REGION Network 9
   RUNG wire#powerrail
      Contact( "I1_7" )
      wire#w1
      Contact( "DB12"."2#回转窑烟气管道闸板上升" )
      I_Contact( "I1_5" )
      I_Contact( "闸阀上限" )
      I_Contact( "Q2_1" )
      Coil( "Q2_0" )
   END_RUNG
   RUNG wire#w1
      Contact( "DB12"."2#回转窑烟气管道闸板下降" )
      I_Contact( "I1_6" )
      I_Contact( "闸阀下限" )
      I_Contact( "Q2_0" )
      Coil( "Q2_1" )
   END_RUNG
   // the same network as SCL:
   "Q2_0" := "I1_7" AND "DB12"."2#回转窑烟气管道闸板上升" AND NOT "I1_5" AND NOT "闸阀上限" AND NOT "Q2_1";
   "Q2_1" := "I1_7" AND "DB12"."2#回转窑烟气管道闸板下降" AND NOT "I1_6" AND NOT "闸阀下限" AND NOT "Q2_0";
END_REGION

REGION Network 10
   RUNG wire#powerrail
      Contact( "DB22".STAT3 )
      Contact( "尾排风机高压远程" )
      Coil( "尾排风机高压合闸驱动" )
   END_RUNG
   // the same network as SCL:
   "尾排风机高压合闸驱动" := "DB22".STAT3 AND "尾排风机高压远程";
END_REGION

REGION Network 11
   RUNG wire#powerrail
      Contact( "DB22".STAT4 )
      Coil( "尾排风机高压分闸驱动" )
   END_RUNG
   // the same network as SCL:
   "尾排风机高压分闸驱动" := "DB22".STAT4;
END_REGION

REGION Network 12
   RUNG wire#powerrail
      Contact( "DB22".STAT5 )
      wire#w1
      Contact( "尾排风机变频远程" )
      Contact( "尾排风机变频待机" )
      I_Contact( "尾排风机变频故障" )
      wire#w2
      I_Contact( "Tag_24" )
      Coil( "尾排风机高压柜变频启动" )
   END_RUNG
   RUNG wire#powerrail
      Contact( "尾排风机高压柜变频启动" )
   END_RUNG wire#w1
   RUNG wire#w2
      S_ODT(T_NO := "Tag_24", TV := S5T#3S, R :=, BI =>, RET_VAL =>)
   END_RUNG
   // the same network as SCL:
   #_w1 := ("DB22".STAT5 OR "尾排风机高压柜变频启动") AND "尾排风机变频远程" AND "尾排风机变频待机" AND NOT "尾排风机变频故障";
   "尾排风机高压柜变频启动" := #_w1 AND NOT "Tag_24";
   #_s5time1 := S_ODT(T_NO := "Tag_24", S := #_w1, TV := S5T#3S);
END_REGION

REGION Network 13
   RUNG wire#powerrail
      Contact( "DB22".STAT6 )
      wire#w1
      Contact( "尾排风机变频远程" )
      wire#w2
      I_Contact( "Tag_25" )
      Coil( "尾排风机高压柜变频停止" )
   END_RUNG
   RUNG wire#powerrail
      Contact( "尾排风机变频故障" )
   END_RUNG wire#w1
   RUNG wire#powerrail
      Contact( "尾排风机高压柜变频停止" )
   END_RUNG wire#w1
   RUNG wire#w2
      S_ODT(T_NO := "Tag_25", TV := S5T#3S, R :=, BI =>, RET_VAL =>)
   END_RUNG
   // the same network as SCL:
   #_w1 := ("DB22".STAT6 OR "尾排风机变频故障" OR "尾排风机高压柜变频停止") AND "尾排风机变频远程";
   "尾排风机高压柜变频停止" := #_w1 AND NOT "Tag_25";
   #_s5time1 := S_ODT(T_NO := "Tag_25", S := #_w1, TV := S5T#3S);
END_REGION
END_FUNCTION

FUNCTION "回转窑模拟量给定" : Void   // FC14, LAD
{ S7_Optimized_Access := 'FALSE' }
VERSION : 0.1
BEGIN

REGION Network 1
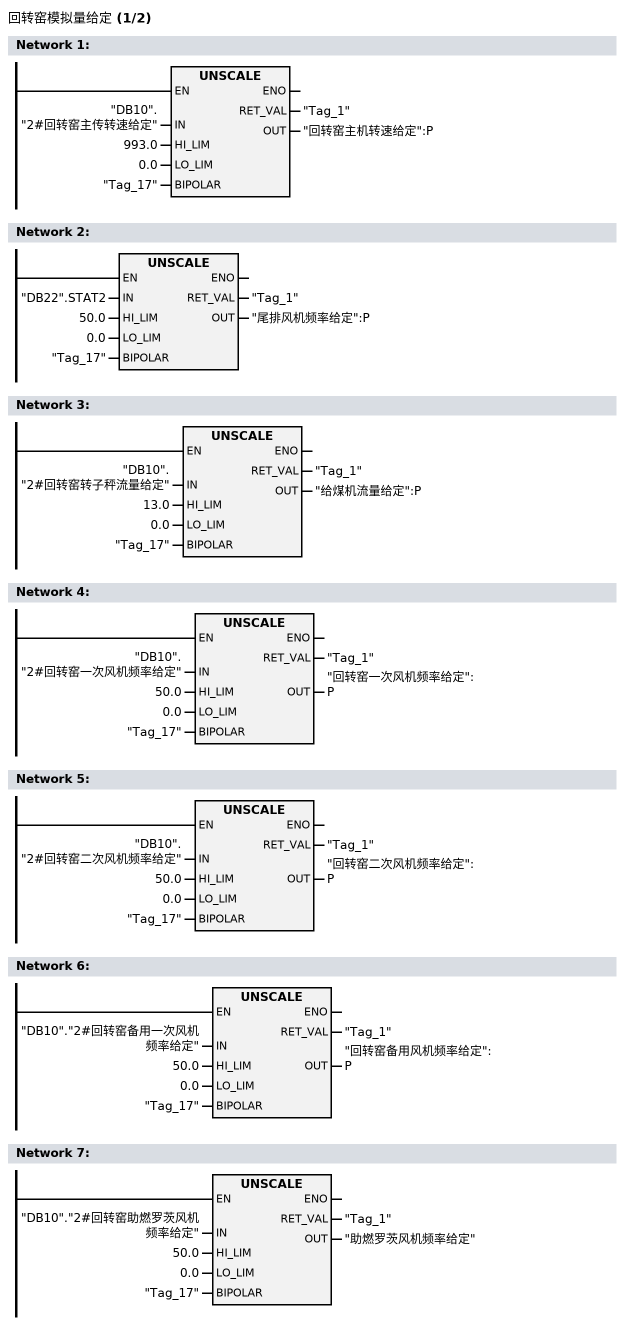
   "Tag_1" := UNSCALE(IN := "DB10"."2#回转窑主传转速给定",
                      HI_LIM := 993.0,
                      LO_LIM := 0.0,
                      BIPOLAR := "Tag_17",
                      OUT => "回转窑主机转速给定":P);
END_REGION

REGION Network 2
   "Tag_1" := UNSCALE(IN := "DB22".STAT2,
                      HI_LIM := 50.0,
                      LO_LIM := 0.0,
                      BIPOLAR := "Tag_17",
                      OUT => "尾排风机频率给定":P);
END_REGION

REGION Network 3
   "Tag_1" := UNSCALE(IN := "DB10"."2#回转窑转子秤流量给定",
                      HI_LIM := 13.0,
                      LO_LIM := 0.0,
                      BIPOLAR := "Tag_17",
                      OUT => "给煤机流量给定":P);
END_REGION

REGION Network 4
   "Tag_1" := UNSCALE(IN := "DB10"."2#回转窑一次风机频率给定",
                      HI_LIM := 50.0,
                      LO_LIM := 0.0,
                      BIPOLAR := "Tag_17",
                      OUT => "回转窑一次风机频率给定":P);
END_REGION

REGION Network 5
   "Tag_1" := UNSCALE(IN := "DB10"."2#回转窑二次风机频率给定",
                      HI_LIM := 50.0,
                      LO_LIM := 0.0,
                      BIPOLAR := "Tag_17",
                      OUT => "回转窑二次风机频率给定":P);
END_REGION

REGION Network 6
   "Tag_1" := UNSCALE(IN := "DB10"."2#回转窑备用一次风机频率给定",
                      HI_LIM := 50.0,
                      LO_LIM := 0.0,
                      BIPOLAR := "Tag_17",
                      OUT => "回转窑备用风机频率给定":P);
END_REGION

REGION Network 7
   "Tag_1" := UNSCALE(IN := "DB10"."2#回转窑助燃罗茨风机频率给定",
                      HI_LIM := 50.0,
                      LO_LIM := 0.0,
                      BIPOLAR := "Tag_17",
                      OUT => "助燃罗茨风机频率给定");
END_REGION

REGION Network 8
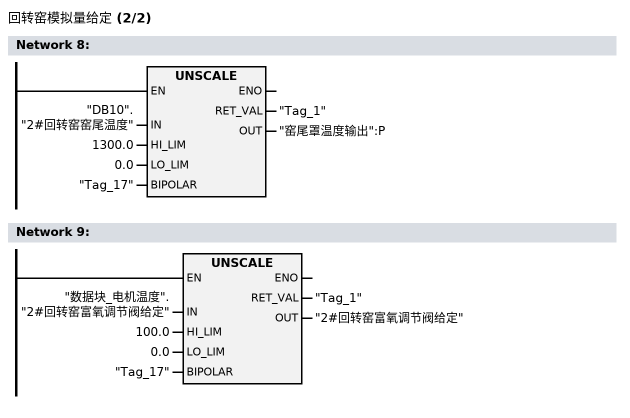
   "Tag_1" := UNSCALE(IN := "DB10"."2#回转窑窑尾温度",
                      HI_LIM := 1300.0,
                      LO_LIM := 0.0,
                      BIPOLAR := "Tag_17",
                      OUT => "窑尾罩温度输出":P);
END_REGION

REGION Network 9
   "Tag_1" := UNSCALE(IN := "数据块_电机温度"."2#回转窑富氧调节阀给定",
                      HI_LIM := 100.0,
                      LO_LIM := 0.0,
                      BIPOLAR := "Tag_17",
                      OUT => "2#回转窑富氧调节阀给定");
END_REGION
END_FUNCTION

FUNCTION "DP&MODBUS通讯" : Void   // FC15, LAD
{ S7_Optimized_Access := 'FALSE' }
VERSION : 0.1
BEGIN

REGION Network 1
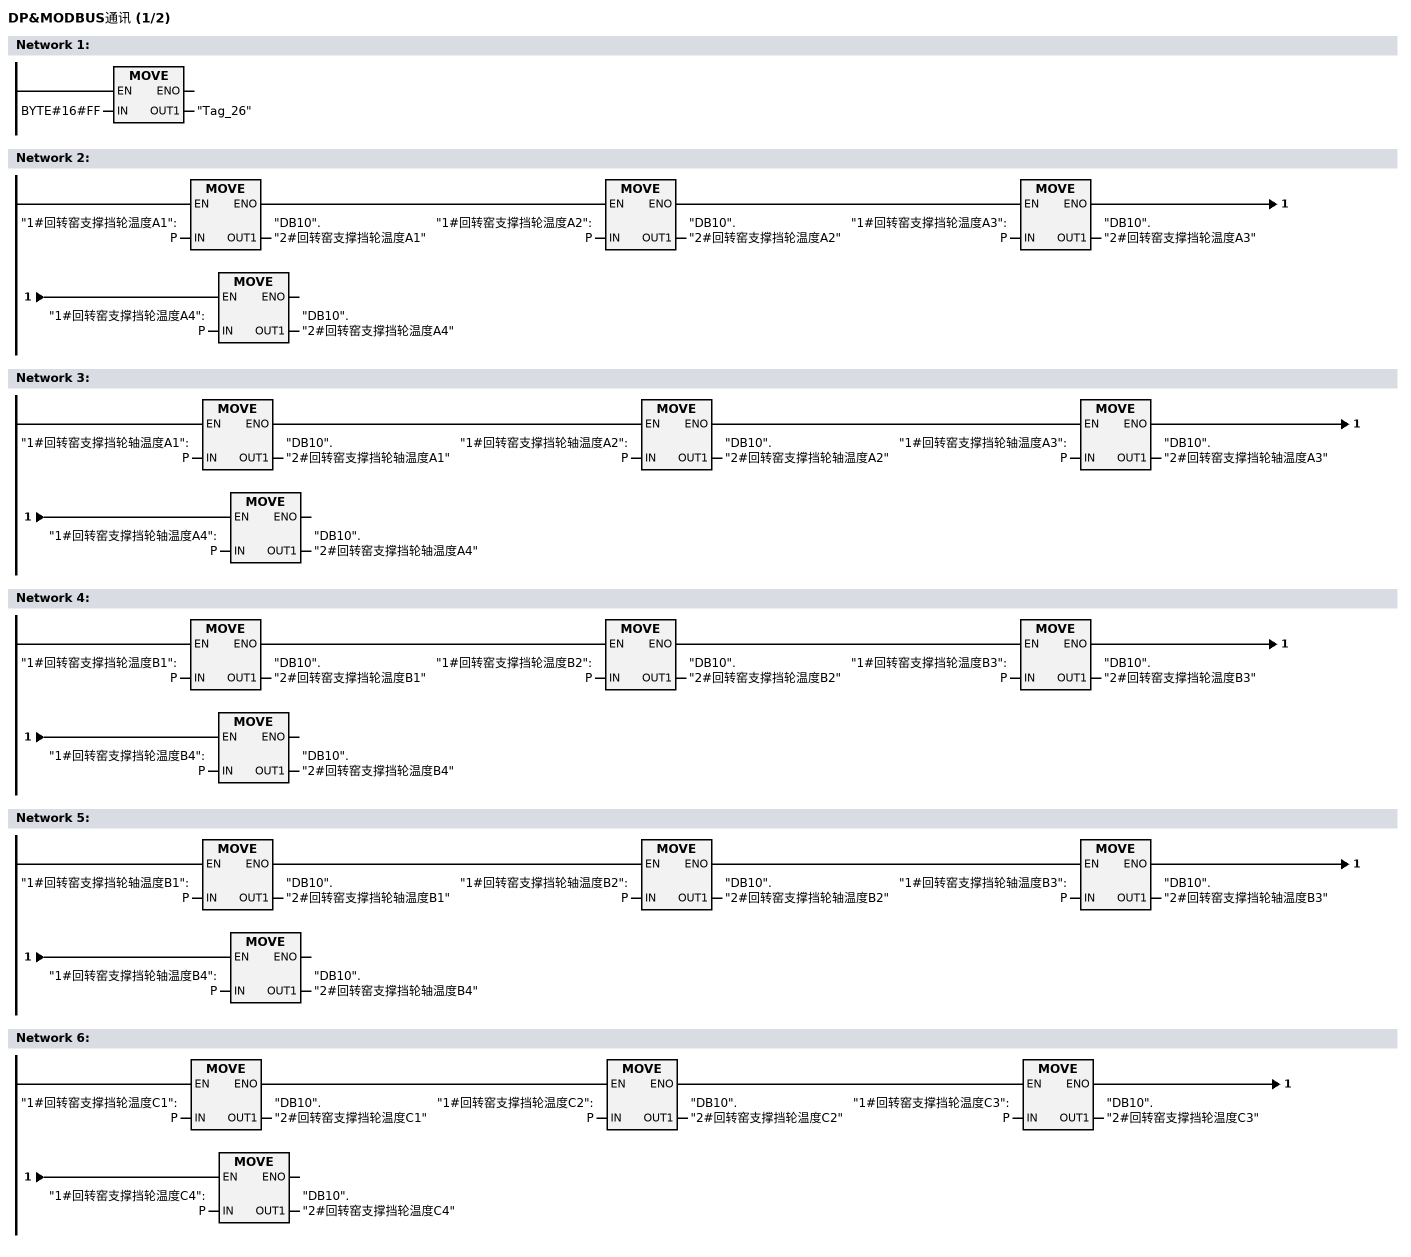
   RUNG wire#powerrail
      { S7_GenerateENO := "TRUE" } Move(in := BYTE#16#FF, out1 => "Tag_26")
   END_RUNG
   // the same network as SCL:
   "Tag_26" := BYTE#16#FF;
END_REGION

REGION Network 2
   RUNG wire#powerrail
      { S7_GenerateENO := "TRUE" } Move(in := "1#回转窑支撑挡轮温度A1":P, out1 => "DB10"."2#回转窑支撑挡轮温度A1")
      { S7_GenerateENO := "TRUE" } Move(in := "1#回转窑支撑挡轮温度A2":P, out1 => "DB10"."2#回转窑支撑挡轮温度A2")
      { S7_GenerateENO := "TRUE" } Move(in := "1#回转窑支撑挡轮温度A3":P, out1 => "DB10"."2#回转窑支撑挡轮温度A3")
      { S7_GenerateENO := "TRUE" } Move(in := "1#回转窑支撑挡轮温度A4":P, out1 => "DB10"."2#回转窑支撑挡轮温度A4")
   END_RUNG
   // the same network as SCL:
   // ENO of a box is taken as its EN; it also drops when the box reports an error
   "DB10"."2#回转窑支撑挡轮温度A1" := "1#回转窑支撑挡轮温度A1":P;
   "DB10"."2#回转窑支撑挡轮温度A2" := "1#回转窑支撑挡轮温度A2":P;
   "DB10"."2#回转窑支撑挡轮温度A3" := "1#回转窑支撑挡轮温度A3":P;
   "DB10"."2#回转窑支撑挡轮温度A4" := "1#回转窑支撑挡轮温度A4":P;
END_REGION

REGION Network 3
   RUNG wire#powerrail
      { S7_GenerateENO := "TRUE" } Move(in := "1#回转窑支撑挡轮轴温度A1":P, out1 => "DB10"."2#回转窑支撑挡轮轴温度A1")
      { S7_GenerateENO := "TRUE" } Move(in := "1#回转窑支撑挡轮轴温度A2":P, out1 => "DB10"."2#回转窑支撑挡轮轴温度A2")
      { S7_GenerateENO := "TRUE" } Move(in := "1#回转窑支撑挡轮轴温度A3":P, out1 => "DB10"."2#回转窑支撑挡轮轴温度A3")
      { S7_GenerateENO := "TRUE" } Move(in := "1#回转窑支撑挡轮轴温度A4":P, out1 => "DB10"."2#回转窑支撑挡轮轴温度A4")
   END_RUNG
   // the same network as SCL:
   // ENO of a box is taken as its EN; it also drops when the box reports an error
   "DB10"."2#回转窑支撑挡轮轴温度A1" := "1#回转窑支撑挡轮轴温度A1":P;
   "DB10"."2#回转窑支撑挡轮轴温度A2" := "1#回转窑支撑挡轮轴温度A2":P;
   "DB10"."2#回转窑支撑挡轮轴温度A3" := "1#回转窑支撑挡轮轴温度A3":P;
   "DB10"."2#回转窑支撑挡轮轴温度A4" := "1#回转窑支撑挡轮轴温度A4":P;
END_REGION

REGION Network 4
   RUNG wire#powerrail
      { S7_GenerateENO := "TRUE" } Move(in := "1#回转窑支撑挡轮温度B1":P, out1 => "DB10"."2#回转窑支撑挡轮温度B1")
      { S7_GenerateENO := "TRUE" } Move(in := "1#回转窑支撑挡轮温度B2":P, out1 => "DB10"."2#回转窑支撑挡轮温度B2")
      { S7_GenerateENO := "TRUE" } Move(in := "1#回转窑支撑挡轮温度B3":P, out1 => "DB10"."2#回转窑支撑挡轮温度B3")
      { S7_GenerateENO := "TRUE" } Move(in := "1#回转窑支撑挡轮温度B4":P, out1 => "DB10"."2#回转窑支撑挡轮温度B4")
   END_RUNG
   // the same network as SCL:
   // ENO of a box is taken as its EN; it also drops when the box reports an error
   "DB10"."2#回转窑支撑挡轮温度B1" := "1#回转窑支撑挡轮温度B1":P;
   "DB10"."2#回转窑支撑挡轮温度B2" := "1#回转窑支撑挡轮温度B2":P;
   "DB10"."2#回转窑支撑挡轮温度B3" := "1#回转窑支撑挡轮温度B3":P;
   "DB10"."2#回转窑支撑挡轮温度B4" := "1#回转窑支撑挡轮温度B4":P;
END_REGION

REGION Network 5
   RUNG wire#powerrail
      { S7_GenerateENO := "TRUE" } Move(in := "1#回转窑支撑挡轮轴温度B1":P, out1 => "DB10"."2#回转窑支撑挡轮轴温度B1")
      { S7_GenerateENO := "TRUE" } Move(in := "1#回转窑支撑挡轮轴温度B2":P, out1 => "DB10"."2#回转窑支撑挡轮轴温度B2")
      { S7_GenerateENO := "TRUE" } Move(in := "1#回转窑支撑挡轮轴温度B3":P, out1 => "DB10"."2#回转窑支撑挡轮轴温度B3")
      { S7_GenerateENO := "TRUE" } Move(in := "1#回转窑支撑挡轮轴温度B4":P, out1 => "DB10"."2#回转窑支撑挡轮轴温度B4")
   END_RUNG
   // the same network as SCL:
   // ENO of a box is taken as its EN; it also drops when the box reports an error
   "DB10"."2#回转窑支撑挡轮轴温度B1" := "1#回转窑支撑挡轮轴温度B1":P;
   "DB10"."2#回转窑支撑挡轮轴温度B2" := "1#回转窑支撑挡轮轴温度B2":P;
   "DB10"."2#回转窑支撑挡轮轴温度B3" := "1#回转窑支撑挡轮轴温度B3":P;
   "DB10"."2#回转窑支撑挡轮轴温度B4" := "1#回转窑支撑挡轮轴温度B4":P;
END_REGION

REGION Network 6
   RUNG wire#powerrail
      { S7_GenerateENO := "TRUE" } Move(in := "1#回转窑支撑挡轮温度C1":P, out1 => "DB10"."2#回转窑支撑挡轮温度C1")
      { S7_GenerateENO := "TRUE" } Move(in := "1#回转窑支撑挡轮温度C2":P, out1 => "DB10"."2#回转窑支撑挡轮温度C2")
      { S7_GenerateENO := "TRUE" } Move(in := "1#回转窑支撑挡轮温度C3":P, out1 => "DB10"."2#回转窑支撑挡轮温度C3")
      { S7_GenerateENO := "TRUE" } Move(in := "1#回转窑支撑挡轮温度C4":P, out1 => "DB10"."2#回转窑支撑挡轮温度C4")
   END_RUNG
   // the same network as SCL:
   // ENO of a box is taken as its EN; it also drops when the box reports an error
   "DB10"."2#回转窑支撑挡轮温度C1" := "1#回转窑支撑挡轮温度C1":P;
   "DB10"."2#回转窑支撑挡轮温度C2" := "1#回转窑支撑挡轮温度C2":P;
   "DB10"."2#回转窑支撑挡轮温度C3" := "1#回转窑支撑挡轮温度C3":P;
   "DB10"."2#回转窑支撑挡轮温度C4" := "1#回转窑支撑挡轮温度C4":P;
END_REGION

REGION Network 7
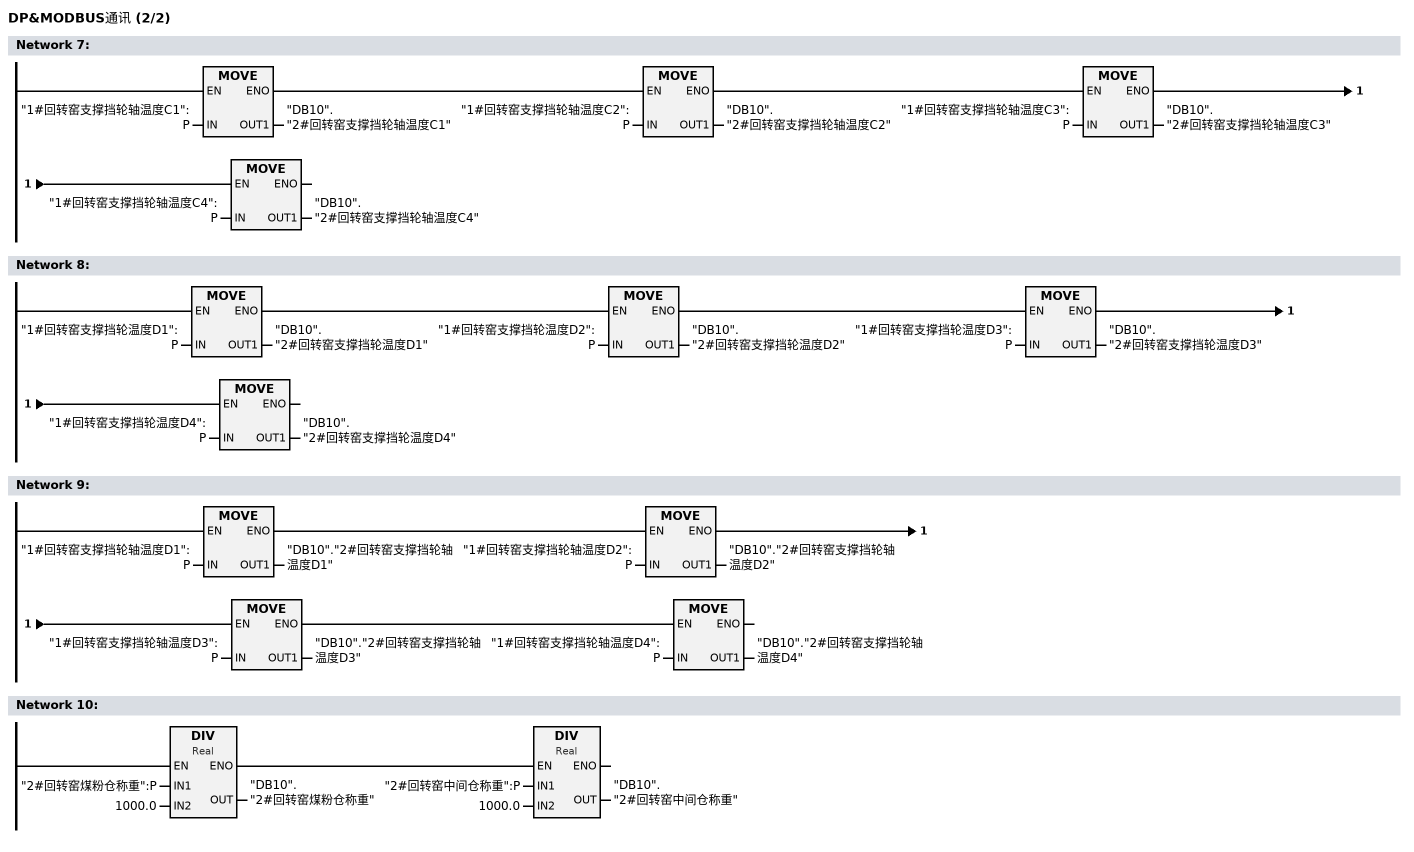
   RUNG wire#powerrail
      { S7_GenerateENO := "TRUE" } Move(in := "1#回转窑支撑挡轮轴温度C1":P, out1 => "DB10"."2#回转窑支撑挡轮轴温度C1")
      { S7_GenerateENO := "TRUE" } Move(in := "1#回转窑支撑挡轮轴温度C2":P, out1 => "DB10"."2#回转窑支撑挡轮轴温度C2")
      { S7_GenerateENO := "TRUE" } Move(in := "1#回转窑支撑挡轮轴温度C3":P, out1 => "DB10"."2#回转窑支撑挡轮轴温度C3")
      { S7_GenerateENO := "TRUE" } Move(in := "1#回转窑支撑挡轮轴温度C4":P, out1 => "DB10"."2#回转窑支撑挡轮轴温度C4")
   END_RUNG
   // the same network as SCL:
   // ENO of a box is taken as its EN; it also drops when the box reports an error
   "DB10"."2#回转窑支撑挡轮轴温度C1" := "1#回转窑支撑挡轮轴温度C1":P;
   "DB10"."2#回转窑支撑挡轮轴温度C2" := "1#回转窑支撑挡轮轴温度C2":P;
   "DB10"."2#回转窑支撑挡轮轴温度C3" := "1#回转窑支撑挡轮轴温度C3":P;
   "DB10"."2#回转窑支撑挡轮轴温度C4" := "1#回转窑支撑挡轮轴温度C4":P;
END_REGION

REGION Network 8
   RUNG wire#powerrail
      { S7_GenerateENO := "TRUE" } Move(in := "1#回转窑支撑挡轮温度D1":P, out1 => "DB10"."2#回转窑支撑挡轮温度D1")
      { S7_GenerateENO := "TRUE" } Move(in := "1#回转窑支撑挡轮温度D2":P, out1 => "DB10"."2#回转窑支撑挡轮温度D2")
      { S7_GenerateENO := "TRUE" } Move(in := "1#回转窑支撑挡轮温度D3":P, out1 => "DB10"."2#回转窑支撑挡轮温度D3")
      { S7_GenerateENO := "TRUE" } Move(in := "1#回转窑支撑挡轮温度D4":P, out1 => "DB10"."2#回转窑支撑挡轮温度D4")
   END_RUNG
   // the same network as SCL:
   // ENO of a box is taken as its EN; it also drops when the box reports an error
   "DB10"."2#回转窑支撑挡轮温度D1" := "1#回转窑支撑挡轮温度D1":P;
   "DB10"."2#回转窑支撑挡轮温度D2" := "1#回转窑支撑挡轮温度D2":P;
   "DB10"."2#回转窑支撑挡轮温度D3" := "1#回转窑支撑挡轮温度D3":P;
   "DB10"."2#回转窑支撑挡轮温度D4" := "1#回转窑支撑挡轮温度D4":P;
END_REGION

REGION Network 9
   RUNG wire#powerrail
      { S7_GenerateENO := "TRUE" } Move(in := "1#回转窑支撑挡轮轴温度D1":P, out1 => "DB10"."2#回转窑支撑挡轮轴温度D1")
      { S7_GenerateENO := "TRUE" } Move(in := "1#回转窑支撑挡轮轴温度D2":P, out1 => "DB10"."2#回转窑支撑挡轮轴温度D2")
      { S7_GenerateENO := "TRUE" } Move(in := "1#回转窑支撑挡轮轴温度D3":P, out1 => "DB10"."2#回转窑支撑挡轮轴温度D3")
      { S7_GenerateENO := "TRUE" } Move(in := "1#回转窑支撑挡轮轴温度D4":P, out1 => "DB10"."2#回转窑支撑挡轮轴温度D4")
   END_RUNG
   // the same network as SCL:
   // ENO of a box is taken as its EN; it also drops when the box reports an error
   "DB10"."2#回转窑支撑挡轮轴温度D1" := "1#回转窑支撑挡轮轴温度D1":P;
   "DB10"."2#回转窑支撑挡轮轴温度D2" := "1#回转窑支撑挡轮轴温度D2":P;
   "DB10"."2#回转窑支撑挡轮轴温度D3" := "1#回转窑支撑挡轮轴温度D3":P;
   "DB10"."2#回转窑支撑挡轮轴温度D4" := "1#回转窑支撑挡轮轴温度D4":P;
END_REGION

REGION Network 10
   RUNG wire#powerrail
      { S7_Templates := "SrcType := Real" } Div(in1 := "2#回转窑煤粉仓称重":P, in2 := 1000.0, out => "DB10"."2#回转窑煤粉仓称重")
      { S7_Templates := "SrcType := Real" } Div(in1 := "2#回转窑中间仓称重":P, in2 := 1000.0, out => "DB10"."2#回转窑中间仓称重")
   END_RUNG
   // the same network as SCL:
   "DB10"."2#回转窑煤粉仓称重" := "2#回转窑煤粉仓称重":P / 1000.0;
   "DB10"."2#回转窑中间仓称重" := "2#回转窑中间仓称重":P / 1000.0;
END_REGION
END_FUNCTION

FUNCTION "配料控制" : Void   // FC21, LAD
{ S7_Optimized_Access := 'FALSE' }
VERSION : 0.1
   VAR_TEMP   // added for the SCL form of the ladder/FBD networks
      _w1 : Bool;
      _w2 : Bool;
   END_VAR
BEGIN

REGION Network 1
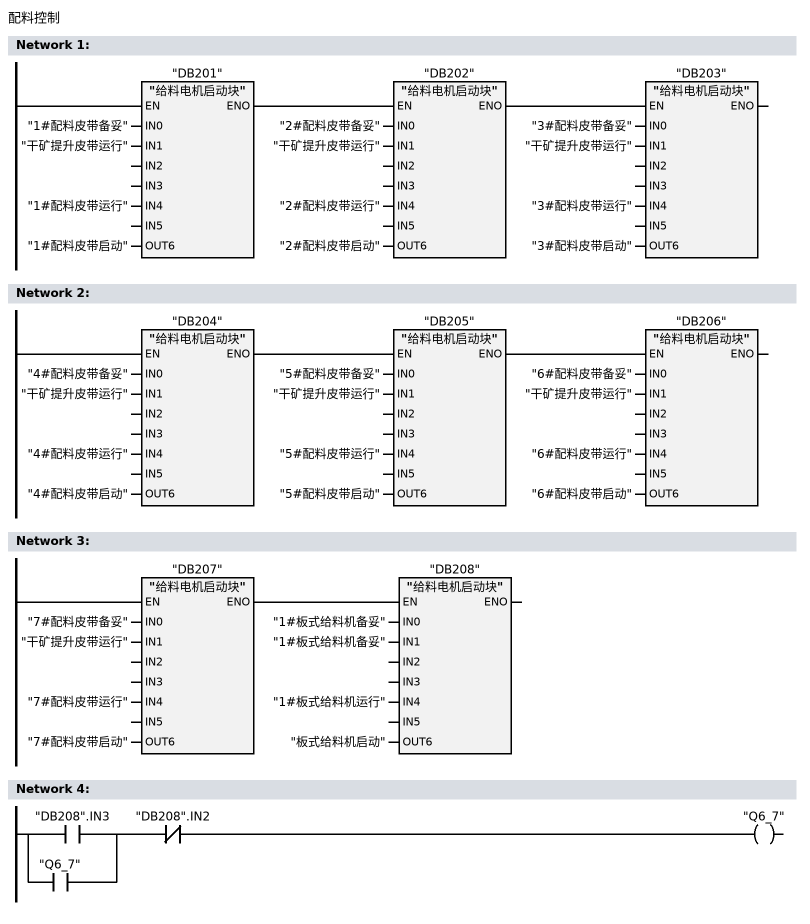
   RUNG wire#powerrail
      "DB201"(IN0 := "1#配料皮带备妥", IN1 := "干矿提升皮带运行", IN2 :=, IN3 :=, IN4 := "1#配料皮带运行", IN5 :=, OUT6 := "1#配料皮带启动")
      "DB202"(IN0 := "2#配料皮带备妥", IN1 := "干矿提升皮带运行", IN2 :=, IN3 :=, IN4 := "2#配料皮带运行", IN5 :=, OUT6 := "2#配料皮带启动")
      "DB203"(IN0 := "3#配料皮带备妥", IN1 := "干矿提升皮带运行", IN2 :=, IN3 :=, IN4 := "3#配料皮带运行", IN5 :=, OUT6 := "3#配料皮带启动")
   END_RUNG
   // the same network as SCL:
   "DB201"(IN0 := "1#配料皮带备妥", IN1 := "干矿提升皮带运行", IN4 := "1#配料皮带运行", OUT6 := "1#配料皮带启动", ENO => #_w1);   // "给料电机启动块"
   "DB202"(EN := #_w1, IN0 := "2#配料皮带备妥", IN1 := "干矿提升皮带运行", IN4 := "2#配料皮带运行", OUT6 := "2#配料皮带启动", ENO => #_w2);   // "给料电机启动块"
   IF #_w2 THEN
       "DB203"(IN0 := "3#配料皮带备妥", IN1 := "干矿提升皮带运行", IN4 := "3#配料皮带运行", OUT6 := "3#配料皮带启动");   // "给料电机启动块"
   END_IF;
END_REGION
